HMI tags "DB_SDC_GLOBAL_REFERENCE"
   "DB_SDC_GLOBAL_REFERENCE_PAR_SET[8].LIMITS" : Array [0..15] of Char = PLC DB_SDC_GLOBAL_REFERENCE.PAR_SET[8].LIMITS AT %DB3786.DBX292.0, 1 s
   "DB_SDC_GLOBAL_REFERENCE_PAR_SET[3].LIMITS" : Array [0..15] of Char = PLC DB_SDC_GLOBAL_REFERENCE.PAR_SET[3].LIMITS AT %DB3786.DBX132.0, 1 s
   "DB_SDC_GLOBAL_REFERENCE_PAR_SET[0].LIMITS" : Array [0..15] of Char = PLC DB_SDC_GLOBAL_REFERENCE.PAR_SET[0].LIMITS AT %DB3786.DBX36.0, 1 s
   "DB_SDC_GLOBAL_REFERENCE_PAR_SET[14].SYNCH" : Array [0..15] of Char = PLC DB_SDC_GLOBAL_REFERENCE.PAR_SET[14].SYNCH AT %DB3786.DBX468.0, 1 s
   "DB_SDC_GLOBAL_REFERENCE_PAR_SET[9].SYNCH" : Array [0..15] of Char = PLC DB_SDC_GLOBAL_REFERENCE.PAR_SET[9].SYNCH AT %DB3786.DBX308.0, 1 s
   "DB_SDC_GLOBAL_REFERENCE_PAR_SET[11].LIMITS" : Array [0..15] of Char = PLC DB_SDC_GLOBAL_REFERENCE.PAR_SET[11].LIMITS AT %DB3786.DBX388.0, 1 s
   "DB_SDC_GLOBAL_REFERENCE_PAR_SET[10].LIMITS" : Array [0..15] of Char = PLC DB_SDC_GLOBAL_REFERENCE.PAR_SET[10].LIMITS AT %DB3786.DBX356.0, 1 s
   "DB_SDC_GLOBAL_REFERENCE_PAR_SET[0].SYNCH" : Array [0..15] of Char = PLC DB_SDC_GLOBAL_REFERENCE.PAR_SET[0].SYNCH AT %DB3786.DBX20.0, 1 s
   "DB_SDC_GLOBAL_REFERENCE_PAR_SET[14].LIMITS" : Array [0..15] of Char = PLC DB_SDC_GLOBAL_REFERENCE.PAR_SET[14].LIMITS AT %DB3786.DBX484.0, 1 s
   "DB_SDC_GLOBAL_REFERENCE_PAR_SET[6].LIMITS" : Array [0..15] of Char = PLC DB_SDC_GLOBAL_REFERENCE.PAR_SET[6].LIMITS AT %DB3786.DBX228.0, 1 s
   "DB_SDC_GLOBAL_REFERENCE_PAR_SET[10].SYNCH" : Array [0..15] of Char = PLC DB_SDC_GLOBAL_REFERENCE.PAR_SET[10].SYNCH AT %DB3786.DBX340.0, 1 s
   "DB_SDC_GLOBAL_REFERENCE_PAR_SET[5].SYNCH" : Array [0..15] of Char = PLC DB_SDC_GLOBAL_REFERENCE.PAR_SET[5].SYNCH AT %DB3786.DBX180.0, 1 s
   "DB_SDC_GLOBAL_REFERENCE_PAR_SET[13].SYNCH" : Array [0..15] of Char = PLC DB_SDC_GLOBAL_REFERENCE.PAR_SET[13].SYNCH AT %DB3786.DBX436.0, 1 s
   "DB_SDC_GLOBAL_REFERENCE_PAR_SET[12].LIMITS" : Array [0..15] of Char = PLC DB_SDC_GLOBAL_REFERENCE.PAR_SET[12].LIMITS AT %DB3786.DBX420.0, 1 s
   "DB_SDC_GLOBAL_REFERENCE_PAR_SET[15].SYNCH" : Array [0..15] of Char = PLC DB_SDC_GLOBAL_REFERENCE.PAR_SET[15].SYNCH AT %DB3786.DBX500.0, 1 s
   "DB_SDC_GLOBAL_REFERENCE_PAR_SET[2].LIMITS" : Array [0..15] of Char = PLC DB_SDC_GLOBAL_REFERENCE.PAR_SET[2].LIMITS AT %DB3786.DBX100.0, 1 s
   "DB_SDC_GLOBAL_REFERENCE_PAR_SET[6].SYNCH" : Array [0..15] of Char = PLC DB_SDC_GLOBAL_REFERENCE.PAR_SET[6].SYNCH AT %DB3786.DBX212.0, 1 s
   "DB_SDC_GLOBAL_REFERENCE_PAR_SET[1].SYNCH" : Array [0..15] of Char = PLC DB_SDC_GLOBAL_REFERENCE.PAR_SET[1].SYNCH AT %DB3786.DBX52.0, 1 s
   "DB_SDC_GLOBAL_REFERENCE_PAR_SET[4].SYNCH" : Array [0..15] of Char = PLC DB_SDC_GLOBAL_REFERENCE.PAR_SET[4].SYNCH AT %DB3786.DBX148.0, 1 s
   "DB_SDC_GLOBAL_REFERENCE_PAR_SET[8].SYNCH" : Array [0..15] of Char = PLC DB_SDC_GLOBAL_REFERENCE.PAR_SET[8].SYNCH AT %DB3786.DBX276.0, 1 s
   "DB_SDC_GLOBAL_REFERENCE_PAR_SET[2].SYNCH" : Array [0..15] of Char = PLC DB_SDC_GLOBAL_REFERENCE.PAR_SET[2].SYNCH AT %DB3786.DBX84.0, 1 s
   "DB_SDC_GLOBAL_REFERENCE_PAR_SET[1].LIMITS" : Array [0..15] of Char = PLC DB_SDC_GLOBAL_REFERENCE.PAR_SET[1].LIMITS AT %DB3786.DBX68.0, 1 s
   "DB_SDC_GLOBAL_REFERENCE_PAR_SET[15].LIMITS" : Array [0..15] of Char = PLC DB_SDC_GLOBAL_REFERENCE.PAR_SET[15].LIMITS AT %DB3786.DBX516.0, 1 s
   "DB_SDC_GLOBAL_REFERENCE_PAR_SET[11].SYNCH" : Array [0..15] of Char = PLC DB_SDC_GLOBAL_REFERENCE.PAR_SET[11].SYNCH AT %DB3786.DBX372.0, 1 s
   "DB_SDC_GLOBAL_REFERENCE_PAR_SET[3].SYNCH" : Array [0..15] of Char = PLC DB_SDC_GLOBAL_REFERENCE.PAR_SET[3].SYNCH AT %DB3786.DBX116.0, 1 s
   "DB_SDC_GLOBAL_REFERENCE_PAR_SET[4].LIMITS" : Array [0..15] of Char = PLC DB_SDC_GLOBAL_REFERENCE.PAR_SET[4].LIMITS AT %DB3786.DBX164.0, 1 s
   "DB_SDC_GLOBAL_REFERENCE_PAR_SET[12].SYNCH" : Array [0..15] of Char = PLC DB_SDC_GLOBAL_REFERENCE.PAR_SET[12].SYNCH AT %DB3786.DBX404.0, 1 s
   "DB_SDC_GLOBAL_REFERENCE_PAR_SET[9].LIMITS" : Array [0..15] of Char = PLC DB_SDC_GLOBAL_REFERENCE.PAR_SET[9].LIMITS AT %DB3786.DBX324.0, 1 s
   "DB_SDC_GLOBAL_REFERENCE_PAR_SET[7].SYNCH" : Array [0..15] of Char = PLC DB_SDC_GLOBAL_REFERENCE.PAR_SET[7].SYNCH AT %DB3786.DBX244.0, 1 s
   "DB_SDC_GLOBAL_REFERENCE_PAR_SET[7].LIMITS" : Array [0..15] of Char = PLC DB_SDC_GLOBAL_REFERENCE.PAR_SET[7].LIMITS AT %DB3786.DBX260.0, 1 s
   "DB_SDC_GLOBAL_REFERENCE_PAR_SET[13].LIMITS" : Array [0..15] of Char = PLC DB_SDC_GLOBAL_REFERENCE.PAR_SET[13].LIMITS AT %DB3786.DBX452.0, 1 s
   "DB_SDC_GLOBAL_REFERENCE_PAR_SET[5].LIMITS" : Array [0..15] of Char = PLC DB_SDC_GLOBAL_REFERENCE.PAR_SET[5].LIMITS AT %DB3786.DBX196.0, 1 s
   "SDC\DB_SDC_GLOBAL_REFERENCE\DB_SDC_GLOBAL_REFERENCE.PROFIL[XX].SORTE" : Array [0..5] of Char AT %DB0.DBX0.0, 1 s
   "DB_SDC_GLOBAL_REFERENCE_HEADER.START_PROFIL" : Int = PLC DB_SDC_GLOBAL_REFERENCE.HEADER.START_PROFIL AT %DB3786.DBW14, 1 s
   "DB_SDC_GLOBAL_REFERENCE_HEADER.LAENGE_PROFIL" : Int = PLC DB_SDC_GLOBAL_REFERENCE.HEADER.LAENGE_PROFIL AT %DB3786.DBW16, 1 s
   "_DB_SDC_GLOBAL_REFERENCE.PROFIL[XX].SORTE_Byte" : Int, internal
   "DB_SDC_GLOBAL_REFERENCE_HEADER.MIN_PROFIL" : Int = PLC DB_SDC_GLOBAL_REFERENCE.HEADER.MIN_PROFIL AT %DB3786.DBW10, 1 s
   "DB_SDC_GLOBAL_REFERENCE_HEADER.MAX_PROFIL" : Int = PLC DB_SDC_GLOBAL_REFERENCE.HEADER.MAX_PROFIL AT %DB3786.DBW12, 1 s
   "_DB_SDC_GLOBAL_REFERENCE.PROFIL[XX+1].SORTE_Byte" : Int, internal
   "SDC\DB_SDC_GLOBAL_REFERENCE\DB_SDC_GLOBAL_REFERENCE.PROFIL[XX+1].SORTE" : Array [0..5] of Char AT %DB0.DBX0.0, 1 s
   "DB_SDC_GLOBAL_REFERENCE_HEADER.DB_NR" : Int = PLC DB_SDC_GLOBAL_REFERENCE.HEADER.DB_NR AT %DB3786.DBW0, 1 s

HMI tags "DB_SDC_EMS_TA"
   "DB_SDC_EMS_TA_HEADER.DB_NR" : Int = PLC DB_SDC_EMS_TA.HEADER.DB_NR AT %DB3728.DBW0, 1 s
   "DB_SDC_EMS_TA_HEADER.MIN_NR_EMS" : Int = PLC DB_SDC_EMS_TA.HEADER.MIN_NR_EMS AT %DB3728.DBW2, 1 s
   "DB_SDC_EMS_TA_HEADER.MAX_NR_EMS" : Int = PLC DB_SDC_EMS_TA.HEADER.MAX_NR_EMS AT %DB3728.DBW4, 1 s
   "DB_SDC_EMS_TA_HEADER.START_EMS" : Int = PLC DB_SDC_EMS_TA.HEADER.START_EMS AT %DB3728.DBW6, 1 s
   "DB_SDC_EMS_TA_HEADER.LAENGE_TA_DATA" : Int = PLC DB_SDC_EMS_TA.HEADER.LAENGE_TA_DATA AT %DB3728.DBW8, 1 s
   "DB_SDC_EMS_TA_HEADER.ANZ_TA" : Int = PLC DB_SDC_EMS_TA.HEADER.ANZ_TA AT %DB3728.DBW10, 1 s
   "DB_SDC_EMS_TA.EMS[XX].TA1.PW1" : Int AT %DB0.DBW0, 1 s
   "_Byte_DB_SDC_EMS_TA.EMS[XX].TA1.PW1" : DInt, internal
   "_Byte_DB_SDC_EMS_TA.EMS[XX].TA1.PW2" : DInt, internal
   "_Byte_DB_SDC_EMS_TA.EMS[XX].TA1.PW3" : DInt, internal
   "_Byte_DB_SDC_EMS_TA.EMS[XX].TA2.PW1" : DInt, internal
   "_Byte_DB_SDC_EMS_TA.EMS[XX].TA2.PW2" : DInt, internal
   "_Byte_DB_SDC_EMS_TA.EMS[XX].TA2.PW3" : DInt, internal
   "_Byte_DB_SDC_EMS_TA.EMS[XX].TA3.PW1" : DInt, internal
   "_Byte_DB_SDC_EMS_TA.EMS[XX].TA3.PW2" : DInt, internal
   "_Byte_DB_SDC_EMS_TA.EMS[XX].TA3.PW3" : DInt, internal
   "DB_SDC_EMS_TA.EMS[XX].TA1.PW2" : Int AT %DB0.DBW0, 1 s
   "DB_SDC_EMS_TA.EMS[XX].TA1.PW3" : Int AT %DB0.DBW0, 1 s
   "DB_SDC_EMS_TA.EMS[XX].TA2.PW1" : Int AT %DB0.DBW0, 1 s
   "DB_SDC_EMS_TA.EMS[XX].TA2.PW2" : Int AT %DB0.DBW0, 1 s
   "DB_SDC_EMS_TA.EMS[XX].TA2.PW3" : Int AT %DB0.DBW0, 1 s
   "DB_SDC_EMS_TA.EMS[XX].TA3.PW1" : Int AT %DB0.DBW0, 1 s
   "DB_SDC_EMS_TA.EMS[XX].TA3.PW2" : Int AT %DB0.DBW0, 1 s
   "DB_SDC_EMS_TA.EMS[XX].TA3.PW3" : Int AT %DB0.DBW0, 1 s
   "DB_SDC_EMS_TA.EMS[XX].TA1.FAULT" : Int AT %DB0.DBW0, 1 s
   "_Byte_DB_SDC_EMS_TA.EMS[XX].TA1.FAULT" : Int AT %MW36, 1 s
   "_Byte_DB_SDC_EMS_TA.EMS[XX].TA1.ALARM" : Int AT %MW38, 1 s
   "_Byte_DB_SDC_EMS_TA.EMS[XX].TA2.FAULT" : DInt, internal
   "_Byte_DB_SDC_EMS_TA.EMS[XX].TA2.ALARM" : DInt, internal
   "_Byte_DB_SDC_EMS_TA.EMS[XX].TA3.FAULT" : DInt, internal
   "_Byte_DB_SDC_EMS_TA.EMS[XX].TA3.ALARM" : DInt, internal
   "DB_SDC_EMS_TA.EMS[XX].TA1.ALARM" : Int AT %DB0.DBW0, 1 s

HMI tags "DB_SDC_TS_IF"
   "DB_SDC_TS_IF_COMMAND_HEADER.DB_NR" : Int = PLC DB_SDC_TS_IF_COMMAND.HEADER.DB_NR AT %DB3716.DBW0, 1 s
   "DB_SDC_TS_IF_COMMAND_HEADER.MIN_NR_SEK" : Int = PLC DB_SDC_TS_IF_COMMAND.HEADER.MIN_NR_SEK AT %DB3716.DBW2, 1 s
   "DB_SDC_TS_IF_COMMAND_HEADER.MAX_NR_SEK" : Int = PLC DB_SDC_TS_IF_COMMAND.HEADER.MAX_NR_SEK AT %DB3716.DBW4, 1 s
   "DB_SDC_TS_IF_COMMAND_HEADER.START_DAT" : Int = PLC DB_SDC_TS_IF_COMMAND.HEADER.START_DAT AT %DB3716.DBW6, 1 s
   "DB_SDC_TS_IF_COMMAND_HEADER.LAENGE_SEK_DATA" : Int = PLC DB_SDC_TS_IF_COMMAND.HEADER.LAENGE_SEK_DATA AT %DB3716.DBW8, 1 s
   "DB_SDC_TS_IF_COMMAND.SEK[XXX].VAL.PROFIL" : Int AT %DB0.DBW0, 1 s
   "_Byte_DB_SDC_TS_IF_COMMAND.SEK[XXX].VAL.PROFIL" : Int, internal
   "DB_SDC_TS_IF_COMMAND_2_HEADER.DB_NR" : Int = PLC DB_SDC_TS_IF_COMMAND_2.HEADER.DB_NR AT %DB3717.DBW0, 1 s
   "DB_SDC_TS_IF_COMMAND_2_HEADER.LAENGE_SEK_DATA" : Int = PLC DB_SDC_TS_IF_COMMAND_2.HEADER.LAENGE_SEK_DATA AT %DB3717.DBW8, 1 s
   "DB_SDC_TS_IF_COMMAND_2_HEADER.MAX_NR_SEK" : Int = PLC DB_SDC_TS_IF_COMMAND_2.HEADER.MAX_NR_SEK AT %DB3717.DBW4, 1 s
   "DB_SDC_TS_IF_COMMAND_2_HEADER.MIN_NR_SEK" : Int = PLC DB_SDC_TS_IF_COMMAND_2.HEADER.MIN_NR_SEK AT %DB3717.DBW2, 1 s
   "DB_SDC_TS_IF_COMMAND_2_HEADER.START_DAT" : Int = PLC DB_SDC_TS_IF_COMMAND_2.HEADER.START_DAT AT %DB3717.DBW6, 1 s
   "_DB_SDC_TS_IF_COMMAND.HEADER.DB_NR" : Int AT %DB716.DBW0
   "_Byte_DB_SDC_TS_IF_COMMAND.SEK[XXX].VAL.D_SETSPEED" : Int, internal
   "DB_SDC_TS_IF_COMMAND.SEK[XXX].VAL.D_SETSPEED" : DInt AT %DB0.DBD0, 1 s
   "_Byte_DB_SDC_TS_IF_COMMAND.SEK[XXX].VAL.D_POS_OFFS" : Int, internal
   "DB_SDC_TS_IF_COMMAND.SEK[XXX].VAL.D_POS_OFFS" : Int AT %DB0.DBW0, 1 s
   "_Byte_DB_SDC_TS_IF_COMMAND.SEK[XXX].BIT1" : Int, internal
   "DB_SDC_TS_IF_COMMAND.SEK[XXX].BIT1" : Int AT %DB0.DBW0, 1 s
   "DB_SDC_TS_IF_COMMAND.SEK[XXX].BIT2" : Int AT %DB0.DBW0, 1 s
   "_Byte_DB_SDC_TS_IF_COMMAND.SEK[XXX].BIT2" : Int, internal
   "DB_SDC_TS_IF_COMMAND.SEK[XXX].BIT3" : Int AT %DB0.DBW0, 1 s
   "_Byte_DB_SDC_TS_IF_COMMAND.SEK[XXX].BIT3" : Int, internal
   "DB_SDC_TS_IF_COMMAND.SEK[XXX].FKT_SET" : Int AT %DB0.DBW0, 1 s
   "_Byte_DB_SDC_TS_IF_COMMAND.SEK[XXX].FKT_SET" : Int, internal
   "DB_SDC_TS_IF_COMMAND.SEK[XXX].FKT_RESET" : Int AT %DB0.DBW0, 1 s
   "_Byte_DB_SDC_TS_IF_COMMAND.SEK[XXX].FKT_RESET" : Int, internal
   "_DB_SDC_TS_IF_STATUS.HEADER.DB_NR" : Int AT %DB716.DBW0
   "_Byte_DB_SDC_TS_IF_STATUS.SEK[XXX].BIT1" : Int, internal
   "_Byte_DB_SDC_TS_IF_STATUS.SEK[XXX].BIT2" : Int, internal
   "_Byte_DB_SDC_TS_IF_STATUS.SEK[XXX].BIT3" : Int, internal
   "_Byte_DB_SDC_TS_IF_STATUS.SEK[XXX].FKT_SET" : Int, internal
   "_Byte_DB_SDC_TS_IF_STATUS.SEK[XXX].VAL.DRIVE_POS" : Int, internal
   "_Byte_DB_SDC_TS_IF_STATUS.SEK[XXX].VAL.PROFIL" : Int, internal
   "_Byte_DB_SDC_TS_IF_STATUS.SEK[XXX].VAL.EMS_ID" : Int, internal
   "DB_SDC_TS_IF_STATUS_HEADER.DB_NR" : Int = PLC DB_SDC_TS_IF_STATUS.HEADER.DB_NR AT %DB3718.DBW0, 1 s
   "DB_SDC_TS_IF_STATUS_HEADER.LAENGE_SEK_DATA" : Int = PLC DB_SDC_TS_IF_STATUS.HEADER.LAENGE_SEK_DATA AT %DB3718.DBW8, 1 s
   "DB_SDC_TS_IF_STATUS_HEADER.MAX_NR_SEK" : Int = PLC DB_SDC_TS_IF_STATUS.HEADER.MAX_NR_SEK AT %DB3718.DBW4, 1 s
   "DB_SDC_TS_IF_STATUS_HEADER.MIN_NR_SEK" : Int = PLC DB_SDC_TS_IF_STATUS.HEADER.MIN_NR_SEK AT %DB3718.DBW2, 1 s
   "DB_SDC_TS_IF_STATUS_HEADER.START_DAT" : Int = PLC DB_SDC_TS_IF_STATUS.HEADER.START_DAT AT %DB3718.DBW6, 1 s
   "DB_SDC_TS_IF_STATUS.SEK[XXX].BIT1" : Int AT %DB0.DBW0, 1 s
   "DB_SDC_TS_IF_STATUS.SEK[XXX].BIT2" : Int AT %DB0.DBW0, 1 s
   "DB_SDC_TS_IF_STATUS.SEK[XXX].BIT3" : Int AT %DB0.DBW0, 1 s
   "DB_SDC_TS_IF_STATUS.SEK[XXX].FKT_SET" : Int AT %DB0.DBW0, 1 s
   "DB_SDC_TS_IF_STATUS.SEK[XXX].VAL.DRIVE_POS" : DInt AT %DB0.DBD0, 1 s
   "DB_SDC_TS_IF_STATUS.SEK[XXX].VAL.PROFIL" : Int AT %DB0.DBW0, 1 s
   "DB_SDC_TS_IF_STATUS.SEK[XXX].VAL.EMS_ID" : Int AT %DB0.DBW0, 1 s
   "DB_SDC_TS_IF_STATUS_2_HEADER.DB_NR" : Int = PLC DB_SDC_TS_IF_STATUS_2.HEADER.DB_NR AT %DB3719.DBW0, 1 s
   "DB_SDC_TS_IF_STATUS_2_HEADER.LAENGE_SEK_DATA" : Int = PLC DB_SDC_TS_IF_STATUS_2.HEADER.LAENGE_SEK_DATA AT %DB3719.DBW8, 1 s
   "DB_SDC_TS_IF_STATUS_2_HEADER.MAX_NR_SEK" : Int = PLC DB_SDC_TS_IF_STATUS_2.HEADER.MAX_NR_SEK AT %DB3719.DBW4, 1 s
   "DB_SDC_TS_IF_STATUS_2_HEADER.MIN_NR_SEK" : Int = PLC DB_SDC_TS_IF_STATUS_2.HEADER.MIN_NR_SEK AT %DB3719.DBW2, 1 s
   "DB_SDC_TS_IF_STATUS_2_HEADER.START_DAT" : Int = PLC DB_SDC_TS_IF_STATUS_2.HEADER.START_DAT AT %DB3719.DBW6, 1 s
   "DB_SDC_TS_IF_STATUS.SEK[XXX].BIT4" : Int AT %DB0.DBW0, 1 s
   "_Byte_DB_SDC_TS_IF_STATUS.SEK[XXX].BIT4" : Int, internal
   "DB_SDC_TS_IF_STATUS.SEK[XXX].SORTE" : Array [0..3] of Char AT %DB0.DBX0.0, 1 s
   "_Byte_DB_SDC_TS_IF_STATUS.SEK[XXX].SORTE" : Int, internal
   "DB_SDC_TS_IF_STATUS.SEK[XXX].VAL.HOIST_POS" : Int AT %DB0.DBW0, 1 s
   "_Byte_DB_SDC_TS_IF_STATUS.SEK[XXX].VAL.HOIST_POS" : Int, internal
   "DB_SDC_TS_IF_STATUS.SEK[XXX].VAL.TILT_POS" : Int AT %DB0.DBW0, 1 s
   "_Byte_DB_SDC_TS_IF_STATUS.SEK[XXX].VAL.TILT_POS" : Int, internal
   "DB_SDC_TS_IF_STATUS.SEK[XXX].VAL.ERROR" : Int AT %DB0.DBW0, 1 s
   "_Byte_DB_SDC_TS_IF_STATUS.SEK[XXX].VAL.ERROR" : Int, internal
   "DB_SDC_TS_IF_STATUS.SEK[XXX].VAL.DRIVE_POS_PERC" : Int AT %DB0.DBW0, 1 s
   "_Byte_DB_SDC_TS_IF_STATUS.SEK[XXX].VAL.DRIVE_POS_PERC" : Int, internal
   "DB_SDC_TS_IF_STATUS.SEK[XXX].VAL.SEK" : Int AT %DB0.DBW0, 1 s
   "_Byte_DB_SDC_TS_IF_STATUS.SEK[XXX].VAL.SEK" : Int, internal
   "DB_SDC_TS_IF_HMI_HEADER.DB_NR" : Int = PLC DB_SDC_TS_IF_HMI.HEADER.DB_NR AT %DB3816.DBW0, 1 s
   "DB_SDC_TS_IF_HMI_HEADER.START_DAT" : Int = PLC DB_SDC_TS_IF_HMI.HEADER.START_DAT AT %DB3816.DBW6, 1 s
   "DB_SDC_TS_IF_HMI_HEADER.LAENGE_SEK_COM" : Int = PLC DB_SDC_TS_IF_HMI.HEADER.LAENGE_SEK_COM AT %DB3816.DBW8, 1 s
   "DB_SDC_TS_IF_HMI_HEADER.LAENGE_SEK_STAT" : Int = PLC DB_SDC_TS_IF_HMI.HEADER.LAENGE_SEK_STAT AT %DB3816.DBW10, 1 s
   "DB_SDC_TS_IF_HMI_HEADER.OFFEST_SEK_STAT" : Int = PLC DB_SDC_TS_IF_HMI.HEADER.OFFEST_SEK_STAT AT %DB3816.DBW12, 1 s
   "DB_SDC_TS_IF_HMI_HEADER.START_HMI" : Int = PLC DB_SDC_TS_IF_HMI.HEADER.START_HMI AT %DB3816.DBW16, 1 s
   "DB_SDC_TS_IF_HMI_HEADER.OFFEST_HMI_DATA" : Int = PLC DB_SDC_TS_IF_HMI.HEADER.OFFEST_HMI_DATA AT %DB3816.DBW18, 1 s
   "_DB_SDC_TS_IF_HMI.HMI_Byte_00" : Int, internal
   "_DB_SDC_TS_IF_HMI.HMI_Byte_02" : Int, internal
   "_DB_SDC_TS_IF_HMI.HMI_Byte_04" : Int, internal
   "_DB_SDC_TS_IF_HMI.HMI_Byte_06" : Int, internal
   "_DB_SDC_TS_IF_HMI.HMI_Byte_08" : Int, internal
   "_DB_SDC_TS_IF_HMI.HMI_Byte_09" : Int, internal
   "_DB_SDC_TS_IF_HMI.HMI_Byte_10" : Int, internal
   "_DB_SDC_TS_IF_HMI.HMI_Byte_12" : Int, internal
   "_DB_SDC_TS_IF_HMI.HMI_Byte_14" : Int, internal
   "_DB_SDC_TS_IF_HMI.HMI_Byte_16" : Int, internal
   "_DB_SDC_TS_IF_HMI.HMI_Byte_18" : Int, internal
   "_DB_SDC_TS_IF_HMI.HMI_Byte_19" : Int, internal
   "DB_SDC_TS_IF_HMI.HMI[XX].BILD_Nr" : Int AT %DB0.DBW0, 1 s   // Bild_Nr aktiv
   "DB_SDC_TS_IF_HMI.HMI[XX].SEK_Nr" : Int AT %DB0.DBW0, 1 s   // Bild_Nr aktiv

HMI tags "DB_SDC_EMS_PAR_ALLG"
   "DB_SDC_EMS_PAR_HMI_HEADER.DB_NR" : Int = PLC DB_SDC_EMS_PAR_HMI.HEADER.DB_NR AT %DB3802.DBW0, 1 s
   "DB_SDC_EMS_PAR_HMI_HEADER.START_PAR" : Int = PLC DB_SDC_EMS_PAR_HMI.HEADER.START_PAR AT %DB3802.DBW6, 1 s
   "DB_SDC_EMS_PAR_HMI_HEADER.LAENGE_PAR" : Int = PLC DB_SDC_EMS_PAR_HMI.HEADER.LAENGE_PAR AT %DB3802.DBW8, 1 s
   "DB_SDC_EMS_PAR_HMI_HMI[1].PULT_Nr_EDIT" : Int = PLC DB_SDC_EMS_PAR_HMI.HMI[1].PULT_Nr_EDIT AT %DB3802.DBW20, 1 s
   "DB_SDC_EMS_PAR_HMI.HMI[XX].BILD_Nr" : Int AT %DB0.DBW0, 1 s
   "DB_SDC_EMS_PAR_HMI.HMI[XX].BILD_Nr_Alt" : Int AT %DB0.DBW0, 1 s
   "_PAR_HMI_Byte_00" : Int, internal
   "_PAR_HMI_Byte_02" : Int, internal
   "_PAR_HMI_Byte_04" : Int, internal
   "_PAR_HMI_Byte_06" : Int, internal
   "_PAR_HMI_Byte_08" : Int, internal
   "_PAR_HMI_Byte_09" : Int, internal
   "_PAR_HMI_Byte_10" : Int, internal
   "_PAR_HMI_Byte_12" : Int, internal
   "_PAR_HMI_Byte_14" : Int, internal
   "_PAR_HMI_Byte_16" : Int, internal
   "_PAR_HMI_Byte_18" : Int, internal
   "_PAR_HMI_Byte_19" : Int, internal
   "DB_SDC_EMS_PAR_HMI.HMI[XX].FR_EDIT" : Bool AT %DB0.DBX0.0, 1 s   // Freigabe Editieren
   "DB_SDC_EMS_PAR_HMI.HMI[XX].PULT_Nr_EDIT" : Int AT %DB0.DBW0, 1 s   // Pult Nr Editieren Aktiv (HMI 1 = Master)
   "DB_SDC_EMS_PAR_HMI.HMI[XX].T_EDIT" : Bool AT %DB0.DBX0.0, 1 s   // Taster Editieren für Pult aktivieren
   "DB_SDC_EMS_PAR_HMI.HMI[XX].T_LOAD" : Bool AT %DB0.DBX0.3, 1 s   // Taster laden
   "DB_SDC_EMS_PAR_HMI.HMI[XX].T_RESET_BED" : Bool AT %DB0.DBX0.1, 1 s   // Taster Reset Bedienfreigabe Pult Nr Bedienung
   "DB_SDC_EMS_PAR_HMI.HMI[XX].T_SAVE" : Bool AT %DB0.DBX0.2, 1 s   // Taster speichern
   "DB_SDC_EMS_PAR_HMI.HMI[XX].ER_DATA" : Bool AT %DB0.DBX0.1, 1 s   // Freigabe Editieren
   "DB_SDC_EMS_PAR_HMI_HEADER.START_HMI" : Int = PLC DB_SDC_EMS_PAR_HMI.HEADER.START_HMI AT %DB3802.DBW16, 1 s
   "DB_SDC_EMS_PAR_HMI_HEADER.OFFEST_HMI_DATA" : Int = PLC DB_SDC_EMS_PAR_HMI.HEADER.OFFEST_HMI_DATA AT %DB3802.DBW18, 1 s

HMI tags "DB_SDC_EMS_PAR_DRIVE"
   "_Byte_EMS[XXX].DRIVE_Delay_Pos" : Int, internal   // Absolute Position / absolute Positon
   "_Byte_EMS[XXX].DRIVE_DelaySpeedContr" : Int, internal   // Absolute Position / absolute Positon
   "_Byte_EMS[XXX].DRIVE_DIV_POS_FAST" : Int, internal   // Absolute Position / absolute Positon
   "_Byte_EMS[XXX].DRIVE_DIV_POS_SLOW" : Int, internal   // Absolute Position / absolute Positon
   "_Byte_EMS[XXX].DRIVE_FUNCT" : Int, internal   // Absolute Position / absolute Positon
   "_Byte_EMS[XXX].DRIVE_TOL_RESET_POS" : Int, internal   // Absolute Position / absolute Positon
   "_Byte_EMS[XXX].DRIVE_TOL_SET_POS" : Int, internal   // Absolute Position / absolute Positon
   "_Byte_EMS[XXX].DRIVE_TolSpeedContr" : Int, internal   // Absolute Position / absolute Positon
   "_Byte_EMS[XXX].DRIVE_V_DIV_FAST" : Int, internal   // Absolute Position / absolute Positon
   "_Byte_EMS[XXX].DRIVE_V_FACT_1" : Int, internal   // Absolute Position / absolute Positon
   "_Byte_EMS[XXX].DRIVE_V_FACT_2" : Int, internal   // Absolute Position / absolute Positon
   "_Byte_EMS[XXX].DRIVE_V_FACT_3" : Int, internal   // Absolute Position / absolute Positon
   "_Byte_EMS[XXX].DRIVE_V_FACT_4" : Int, internal   // Absolute Position / absolute Positon
   "_Byte_EMS[XXX].DRIVE_V_FACT_5" : Int, internal   // Absolute Position / absolute Positon
   "_Byte_EMS[XXX].DRIVE_V_Fixed_1" : Int, internal   // Absolute Position / absolute Positon
   "_Byte_EMS[XXX].DRIVE_V_Fixed_2" : Int, internal   // Absolute Position / absolute Positon
   "_Byte_EMS[XXX].DRIVE_V_Fixed_4_SLS_SPEED" : Int, internal   // Absolute Position / absolute Positon
   "_Byte_EMS[XXX].DRIVE_V_LIMIT_FACT" : Int, internal   // Absolute Position / absolute Positon
   "_Byte_EMS[XXX].DRIVE_V_max_Not_top" : Int, internal   // Absolute Position / absolute Positon
   "_Byte_EMS[XXX].DRIVE_V_max_top" : Int, internal   // Absolute Position / absolute Positon
   "_Byte_EMS[XXX].DRIVE_V_min" : Int, internal   // Absolute Position / absolute Positon
   "_Byte_EMS[XXX].DRIVE_V_Pos_2" : Int, internal   // Absolute Position / absolute Positon
   "_Byte_EMS[XXX].DRIVE_V_SETP_1" : Int, internal   // Absolute Position / absolute Positon
   "_Byte_EMS[XXX].DRIVE_V_SETP_2" : Int, internal   // Absolute Position / absolute Positon
   "_Byte_EMS[XXX].DRIVE_V_SETP_3" : Int, internal   // Absolute Position / absolute Positon
   "_Byte_EMS[XXX].DRIVE_V_SETP_4" : Int, internal   // Absolute Position / absolute Positon
   "_Byte_EMS[XXX].DRIVE_Window_Movement" : Int, internal   // Absolute Position / absolute Positon
   "_Byte_EMS[XXX].DRIVE_Window_Overrun" : Int, internal   // Absolute Position / absolute Positon
   "_Byte_EMS[XXX].DRIVE_Window_Pos" : Int, internal   // Absolute Position / absolute Positon
   "_Byte_EMS[XXX].DRIVE_Window_Pos_2" : Int, internal   // Absolute Position / absolute Positon
   "DB_SDC_EMS_PAR_HMI.HMI[XX].PAR.DRIVE.Delay_Pos" : Int AT %DB0.DBW0, 1 s
   "DB_SDC_EMS_PAR_HMI.HMI[XX].PAR.DRIVE.DelaySpeedContr" : S5Time AT %DB0.DBW0, 1 s
   "DB_SDC_EMS_PAR_HMI.HMI[XX].PAR.DRIVE.DIV_POS_FAST" : DInt AT %DB0.DBD0, 1 s
   "DB_SDC_EMS_PAR_HMI.HMI[XX].PAR.DRIVE.DIV_POS_SLOW" : DInt AT %DB0.DBD0, 1 s
   "DB_SDC_EMS_PAR_HMI.HMI[XX].PAR.DRIVE.TOL_RESET_POS" : Int AT %DB0.DBW0, 1 s
   "DB_SDC_EMS_PAR_HMI.HMI[XX].PAR.DRIVE.TOL_SET_POS" : Int AT %DB0.DBW0, 1 s
   "DB_SDC_EMS_PAR_HMI.HMI[XX].PAR.DRIVE.TolSpeedContr" : Int AT %DB0.DBW0, 1 s
   "DB_SDC_EMS_PAR_HMI.HMI[XX].PAR.DRIVE.V_DIV_FAST" : DInt AT %DB0.DBD0, 1 s
   "DB_SDC_EMS_PAR_HMI.HMI[XX].PAR.DRIVE.V_Fixed_1" : DInt AT %DB0.DBD0, 1 s
   "DB_SDC_EMS_PAR_HMI.HMI[XX].PAR.DRIVE.V_Fixed_2" : DInt AT %DB0.DBD0, 1 s
   "DB_SDC_EMS_PAR_HMI.HMI[XX].PAR.DRIVE.V_Fixed_4_SLS_SPEED" : DInt AT %DB0.DBD0, 1 s
   "DB_SDC_EMS_PAR_HMI.HMI[XX].PAR.DRIVE.V_max_Not_top" : DInt AT %DB0.DBD0, 1 s
   "DB_SDC_EMS_PAR_HMI.HMI[XX].PAR.DRIVE.V_max_top" : DInt AT %DB0.DBD0, 1 s
   "DB_SDC_EMS_PAR_HMI.HMI[XX].PAR.DRIVE.V_min" : DInt AT %DB0.DBD0, 1 s
   "DB_SDC_EMS_PAR_HMI.HMI[XX].PAR.DRIVE.V_Pos_2" : DInt AT %DB0.DBD0, 1 s
   "DB_SDC_EMS_PAR_HMI.HMI[XX].PAR.DRIVE.Window_Movement" : Int AT %DB0.DBW0, 1 s
   "DB_SDC_EMS_PAR_HMI.HMI[XX].PAR.DRIVE.Window_Overrun" : Int AT %DB0.DBW0, 1 s
   "DB_SDC_EMS_PAR_HMI.HMI[XX].PAR.DRIVE.Window_Pos" : Int AT %DB0.DBW0, 1 s
   "DB_SDC_EMS_PAR_HMI.HMI[XX].PAR.DRIVE.Window_Pos_2" : Int AT %DB0.DBW0, 1 s
   "DB_SDC_EMS_PAR_HMI.HMI[XX].PAR.DRIVE.Funct" : Word AT %DB0.DBW0, 1 s
   "DB_SDC_EMS_PAR_HMI.HMI[XX].PAR.DRIVE.V_FACT_1" : Real AT %DB0.DBD0, 1 s
   "DB_SDC_EMS_PAR_HMI.HMI[XX].PAR.DRIVE.V_FACT_2" : Real AT %DB0.DBD0, 1 s
   "DB_SDC_EMS_PAR_HMI.HMI[XX].PAR.DRIVE.V_FACT_3" : Real AT %DB0.DBD0, 1 s
   "DB_SDC_EMS_PAR_HMI.HMI[XX].PAR.DRIVE.V_FACT_4" : Real AT %DB0.DBD0, 1 s
   "DB_SDC_EMS_PAR_HMI.HMI[XX].PAR.DRIVE.V_FACT_5" : Real AT %DB0.DBD0, 1 s
   "DB_SDC_EMS_PAR_HMI.HMI[XX].PAR.DRIVE.V_LIMIT_FACT" : Real AT %DB0.DBD0, 1 s
   "DB_SDC_EMS_PAR_HMI.HMI[XX].PAR.DRIVE.V_SETP_1" : DInt AT %DB0.DBD0, 1 s
   "DB_SDC_EMS_PAR_HMI.HMI[XX].PAR.DRIVE.V_SETP_2" : DInt AT %DB0.DBD0, 1 s
   "DB_SDC_EMS_PAR_HMI.HMI[XX].PAR.DRIVE.V_SETP_3" : DInt AT %DB0.DBD0, 1 s
   "DB_SDC_EMS_PAR_HMI.HMI[XX].PAR.DRIVE.V_SETP_4" : DInt AT %DB0.DBD0, 1 s
   "_Byte_EMS[XXX].DRIVE_Delay_Pos(1)" : Int, internal

HMI tags "DB_SDC_EMS_PAR_HOIST"
   "_Byte_EMS[XXX].HOIST_V_min" : Int, internal   // Absolute Position / absolute Positon
   "DB_SDC_EMS_PAR_HMI.HMI[XX].PAR.HOIST.V_min" : Int AT %DB0.DBW0, 1 s
   "_Byte_EMS[XXX].HOIST_V_max" : Int, internal   // Absolute Position / absolute Positon
   "DB_SDC_EMS_PAR_HMI.HMI[XX].PAR.HOIST.V_max" : Int AT %DB0.DBW0, 1 s
   "_Byte_EMS[XXX].HOIST_V_MaxOccLift" : Int, internal   // Absolute Position / absolute Positon
   "DB_SDC_EMS_PAR_HMI.HMI[XX].PAR.HOIST.V_MaxOccLift" : Int AT %DB0.DBW0, 1 s
   "_Byte_EMS[XXX].HOIST_V_Pos_1" : Int, internal   // Absolute Position / absolute Positon
   "DB_SDC_EMS_PAR_HMI.HMI[XX].PAR.HOIST.V_Pos_1" : Int AT %DB0.DBW0, 1 s
   "_Byte_EMS[XXX].HOIST_V_Pos_2" : Int, internal   // Absolute Position / absolute Positon
   "DB_SDC_EMS_PAR_HMI.HMI[XX].PAR.HOIST.V_Pos_2" : Int AT %DB0.DBW0, 1 s
   "_Byte_EMS[XXX].HOIST_V_Fixed_1" : Int, internal   // Absolute Position / absolute Positon
   "DB_SDC_EMS_PAR_HMI.HMI[XX].PAR.HOIST.V_Fixed_1" : Int AT %DB0.DBW0, 1 s
   "_Byte_EMS[XXX].HOIST_V_Fixed_2" : Int, internal   // Absolute Position / absolute Positon
   "DB_SDC_EMS_PAR_HMI.HMI[XX].PAR.HOIST.V_Fixed_2" : Int AT %DB0.DBW0, 1 s
   "_Byte_EMS[XXX].HOIST_V_Fixed_4" : Int, internal   // Absolute Position / absolute Positon
   "DB_SDC_EMS_PAR_HMI.HMI[XX].PAR.HOIST.V_Fixed_4" : Int AT %DB0.DBW0, 1 s
   "_Byte_EMS[XXX].HOIST_V_Fixed_6" : Int, internal   // Absolute Position / absolute Positon
   "DB_SDC_EMS_PAR_HMI.HMI[XX].PAR.HOIST.V_Fixed_6" : Int AT %DB0.DBW0, 1 s
   "_Byte_EMS[XXX].HOIST_V_FACT_Hz_UP" : Int, internal   // Absolute Position / absolute Positon
   "DB_SDC_EMS_PAR_HMI.HMI[XX].PAR.HOIST.V_FACT_Hz_UP" : Real AT %DB0.DBD0, 1 s
   "_Byte_EMS[XXX].HOIST_V_FACT_Hz_DOWN" : Int, internal   // Absolute Position / absolute Positon
   "DB_SDC_EMS_PAR_HMI.HMI[XX].PAR.HOIST.V_FACT_Hz_DOWN" : Real AT %DB0.DBD0, 1 s
   "DB_SDC_EMS_PAR_HMI.HMI[XX].PAR.HOIST.H_Window_POS_V1" : Int AT %DB0.DBW0, 1 s
   "_Byte_EMS[XXX].HOIST_H_Window_POS_V1" : Int, internal   // Absolute Position / absolute Positon
   "DB_SDC_EMS_PAR_HMI.HMI[XX].PAR.HOIST.H_Window_POS_V2" : Int AT %DB0.DBW0, 1 s
   "_Byte_EMS[XXX].HOIST_H_Window_POS_V2" : Int, internal   // Absolute Position / absolute Positon
   "DB_SDC_EMS_PAR_HMI.HMI[XX].PAR.HOIST.H_TOL_SET_POS" : Int AT %DB0.DBW0, 1 s
   "_Byte_EMS[XXX].HOIST_H_TOL_SET_POS" : Int, internal   // Absolute Position / absolute Positon
   "DB_SDC_EMS_PAR_HMI.HMI[XX].PAR.HOIST.H_TOL_RESET_POS" : Int AT %DB0.DBW0, 1 s
   "_Byte_EMS[XXX].HOIST_H_TOL_RESET_POS" : Int, internal   // Absolute Position / absolute Positon
   "DB_SDC_EMS_PAR_HMI.HMI[XX].PAR.HOIST.H_MIN" : Int AT %DB0.DBW0, 1 s
   "_Byte_EMS[XXX].HOIST_H_MIN" : Int, internal   // Absolute Position / absolute Positon
   "DB_SDC_EMS_PAR_HMI.HMI[XX].PAR.HOIST.H_MIN_without_bypass" : Int AT %DB0.DBW0, 1 s
   "_Byte_EMS[XXX].HOIST_H_MIN_without_bypass" : Int, internal   // Absolute Position / absolute Positon
   "DB_SDC_EMS_PAR_HMI.HMI[XX].PAR.HOIST.H_REF_OFFSET" : Int AT %DB0.DBW0, 1 s
   "_Byte_EMS[XXX].HOIST_H_REF_OFFSET" : Int, internal   // Absolute Position / absolute Positon
   "DB_SDC_EMS_PAR_HMI.HMI[XX].PAR.HOIST.H_REF" : Int AT %DB0.DBW0, 1 s
   "_Byte_EMS[XXX].HOIST_H_REF" : Int, internal   // Absolute Position / absolute Positon
   "DB_SDC_EMS_PAR_HMI.HMI[XX].PAR.HOIST.H_FACT_ENC1" : Real AT %DB0.DBD0, 1 s
   "_Byte_EMS[XXX].HOIST_H_FACT_ENC1" : Int, internal   // Absolute Position / absolute Positon
   "DB_SDC_EMS_PAR_HMI.HMI[XX].PAR.HOIST.H_FACT_ENC2" : Real AT %DB0.DBD0, 1 s
   "_Byte_EMS[XXX].HOIST_H_FACT_ENC2" : Int, internal   // Absolute Position / absolute Positon
   "DB_SDC_EMS_PAR_HMI.HMI[XX].PAR.HOIST.H_FACT_SPEED" : Real AT %DB0.DBD0, 1 s
   "_Byte_EMS[XXX].HOIST_H_FACT_SPEED" : Int, internal   // Absolute Position / absolute Positon
   "DB_SDC_EMS_PAR_HMI.HMI[XX].PAR.HOIST.H_ENC_MAX_DIFF" : Int AT %DB0.DBW0, 1 s
   "_Byte_EMS[XXX].HOIST_H_ENC_MAX_DIFF" : Int, internal   // Absolute Position / absolute Positon
   "DB_SDC_EMS_PAR_HMI.HMI[XX].PAR.HOIST.H_Slow" : Int AT %DB0.DBW0, 1 s
   "_Byte_EMS[XXX].HOIST_H_Slow" : Int, internal   // Absolute Position / absolute Positon
   "DB_SDC_EMS_PAR_HMI.HMI[XX].PAR.HOIST.H_tIN_POS" : Int AT %DB0.DBW0, 1 s
   "_Byte_EMS[XXX].HOIST_H_tIN_POS" : Int, internal   // Absolute Position / absolute Positon
   "DB_SDC_EMS_PAR_HMI.HMI[XX].PAR.HOIST.H_REF_HMI" : Int AT %DB0.DBW0, 1 s
   "_Byte_EMS[XXX].HOIST_H_REF_HMI" : Int, internal   // Absolute Position / absolute Positon
   "_Byte_EMS[XXX].HOIST_V_Fixed_3" : Int, internal
   "DB_SDC_EMS_PAR_HMI.HMI[XX].PAR.HOIST.V_Fixed_3" : Int AT %DB0.DBW0, 1 s

HMI tags "VAT_SYSTEM_ALLG"
   "_intern_BILD_Nr" : Int, internal
   "_intern_1_bool" : Bool, internal
   "_intern_0_bool" : Bool, internal
   "_intern_1" : Int, internal
   "_intern_2" : Int, internal
   "_intern_3" : Int, internal
   "_intern_4" : Int, internal
   "_intern_5" : Int, internal
   "_intern_6" : Int, internal
   "_intern_7" : Int, internal
   "_intern_8" : Int, internal
   "_intern_9" : Int, internal
   "_intern_10" : Int, internal
   "_intern_11" : Int, internal
   "_intern_12" : Int, internal
   "_intern_13" : Int, internal
   "_intern_14" : Int, internal
   "_intern_15" : Int, internal
   "_intern_16" : Int, internal
   "_intern_17" : Int, internal
   "_intern_18" : Int, internal
   "_intern_19" : Int, internal
   "_intern_20" : Int, internal
   "_intern_21" : Int, internal
   "_intern_22" : Int, internal
   "_intern_23" : Int, internal
   "_intern_24" : Int, internal
   "_intern_25" : Int, internal
   "_intern_26" : Int, internal
   "_intern_27" : Int, internal
   "_intern_28" : Int, internal
   "_intern_29" : Int, internal
   "_intern_30" : Int, internal
   "_intern_31" : Int, internal
   "_intern_32" : Int, internal
   "_intern_33" : Int, internal
   "_intern_34" : Int, internal
   "_intern_35" : Int, internal
   "_intern_36" : Int, internal
   "_intern_37" : Int, internal
   "_intern_38" : Int, internal
   "_intern_39" : Int, internal
   "_intern_40" : Int, internal
   "_intern_41" : Int, internal
   "_intern_42" : Int, internal
   "_intern_43" : Int, internal
   "_intern_44" : Int, internal
   "_intern_45" : Int, internal
   "_intern_46" : Int, internal
   "_intern_47" : Int, internal
   "_intern_48" : Int, internal
   "_intern_49" : Int, internal
   "_intern_50" : Int, internal
   "_intern_51" : Int, internal
   "_intern_52" : Int, internal
   "_intern_53" : Int, internal
   "_intern_54" : Int, internal
   "_intern_55" : Int, internal
   "_intern_56" : Int, internal
   "_intern_57" : Int, internal
   "_intern_58" : Int, internal
   "_intern_59" : Int, internal
   "_intern_60" : Int, internal
   "_intern_61" : Int, internal
   "_intern_62" : Int, internal
   "_intern_63" : Int, internal
   "_intern_64" : Int, internal
   "_intern_65" : Int, internal
   "_intern_66" : Int, internal
   "_intern_67" : Int, internal
   "_intern_68" : Int, internal
   "_intern_69" : Int, internal
   "_intern_70" : Int, internal
   "_intern_71" : Int, internal
   "_intern_72" : Int, internal
   "_intern_73" : Int, internal
   "_intern_74" : Int, internal
   "_intern_75" : Int, internal
   "_intern_76" : Int, internal
   "_intern_77" : Int, internal
   "_intern_78" : Int, internal
   "_intern_79" : Int, internal
   "_intern_80" : Int, internal
   "_intern_81" : Int, internal
   "_intern_82" : Int, internal
   "_intern_83" : Int, internal
   "_intern_84" : Int, internal
   "_intern_85" : Int, internal
   "_intern_86" : Int, internal
   "_intern_87" : Int, internal
   "_intern_88" : Int, internal
   "_intern_89" : Int, internal
   "_intern_90" : Int, internal
   "_intern_91" : Int, internal
   "_intern_92" : Int, internal
   "_intern_93" : Int, internal
   "_intern_94" : Int, internal
   "_intern_95" : Int, internal
   "_intern_96" : Int, internal
   "_intern_97" : Int, internal
   "_intern_98" : Int, internal
   "_intern_99" : Int, internal
   "_intern_100" : Int, internal
   "_intern_101" : Int, internal
   "_intern_102" : Int, internal
   "_intern_103" : Int, internal
   "_intern_104" : Int, internal
   "_intern_105" : Int, internal
   "_intern_106" : Int, internal
   "_intern_107" : Int, internal
   "_intern_108" : Int, internal
   "_intern_109" : Int, internal
   "_intern_110" : Int, internal
   "_intern_111" : Int, internal
   "_intern_112" : Int, internal
   "_intern_113" : Int, internal
   "_intern_114" : Int, internal
   "_intern_115" : Int, internal
   "_intern_116" : Int, internal
   "_intern_117" : Int, internal
   "_intern_118" : Int, internal
   "_intern_119" : Int, internal
   "_intern_120" : Int, internal
   "_intern_121" : Int, internal
   "_intern_122" : Int, internal
   "_intern_123" : Int, internal
   "_intern_124" : Int, internal
   "_intern_125" : Int, internal
   "_intern_126" : Int, internal
   "_intern_127" : Int, internal
   "_intern_128" : Int, internal
   "_intern_129" : Int, internal
   "_intern_130" : Int, internal
   "_intern_131" : Int, internal
   "_intern_132" : Int, internal
   "_intern_133" : Int, internal
   "_intern_134" : Int, internal
   "_intern_135" : Int, internal
   "_intern_136" : Int, internal
   "_intern_137" : Int, internal
   "_intern_138" : Int, internal
   "_intern_139" : Int, internal
   "_intern_140" : Int, internal
   "_intern_141" : Int, internal
   "_intern_142" : Int, internal
   "_intern_143" : Int, internal
   "_intern_144" : Int, internal
   "_intern_145" : Int, internal
   "_intern_146" : Int, internal
   "_intern_147" : Int, internal
   "_intern_148" : Int, internal
   "_intern_149" : Int, internal
   "_intern_150" : Int, internal
   "_intern_151" : Int, internal
   "_intern_152" : Int, internal
   "_intern_153" : Int, internal
   "_intern_154" : Int, internal
   "_intern_155" : Int, internal
   "_intern_156" : Int, internal
   "_intern_157" : Int, internal
   "_intern_158" : Int, internal
   "_intern_159" : Int, internal
   "_intern_160" : Int, internal
   "_intern_161" : Int, internal
   "_intern_162" : Int, internal
   "_intern_163" : Int, internal
   "_intern_164" : Int, internal
   "_intern_165" : Int, internal
   "_intern_166" : Int, internal
   "_intern_167" : Int, internal
   "_intern_168" : Int, internal
   "_intern_169" : Int, internal
   "_intern_170" : Int, internal
   "_intern_171" : Int, internal
   "_intern_172" : Int, internal
   "_intern_173" : Int, internal
   "_intern_174" : Int, internal
   "_intern_175" : Int, internal
   "_intern_176" : Int, internal
   "_intern_177" : Int, internal
   "_intern_178" : Int, internal
   "_intern_179" : Int, internal
   "_intern_180" : Int, internal
   "_intern_181" : Int, internal
   "_intern_182" : Int, internal
   "_intern_183" : Int, internal
   "_intern_184" : Int, internal
   "_intern_185" : Int, internal
   "_intern_186" : Int, internal
   "_intern_187" : Int, internal
   "_intern_188" : Int, internal
   "_intern_189" : Int, internal
   "_intern_190" : Int, internal
   "_intern_191" : Int, internal
   "_intern_192" : Int, internal
   "_intern_193" : Int, internal
   "_intern_194" : Int, internal
   "_intern_195" : Int, internal
   "_intern_196" : Int, internal
   "_intern_197" : Int, internal
   "_intern_198" : Int, internal
   "_intern_199" : Int, internal
   "_intern_200" : Int, internal

